REGION Network 2: ADDRESS 2
   RUNG wire#powerrail
      { S7_Templates := "SrcType := Real"; S7_GenerateENO := "TRUE" } Div(in1 := "DB6_MAV2_DBD".ADDRES_2, in2 := 32.768, out => "DB6_MAV2_DBD".SCALLING_2)
      { S7_Templates := "[SrcType := Real, DestType := DInt]"; S7_GenerateENO := "TRUE" } Round(in := "DB6_MAV2_DBD".SCALLING_2, out => "DB6_MAV2_DBD".STAT58)
      { S7_GenerateENO := "TRUE" } Move(in := "DB6_MAV2_DBD".STAT58, out1 => "DB7".STAT0)
   END_RUNG
   // the same network as SCL:
   // ENO of a box is taken as its EN; it also drops when the box reports an error
   "DB6_MAV2_DBD".SCALLING_2 := "DB6_MAV2_DBD".ADDRES_2 / 32.768;
   "DB6_MAV2_DBD".STAT58 := ROUND("DB6_MAV2_DBD".SCALLING_2);
   "DB7".STAT0 := "DB6_MAV2_DBD".STAT58;
END_REGION

REGION Network 3: ADDRESS 3
   RUNG wire#powerrail
      { S7_Templates := "[SrcType := Int, DestType := DInt]"; S7_GenerateENO := "TRUE" } Convert(in := "DB5_MAV".ADDRES_3, out => "DB8_SCALLING_MAV".ADDRESS_3)
      { S7_Templates := "[SrcType := DInt, DestType := Real]"; S7_GenerateENO := "TRUE" } Convert(in := "DB8_SCALLING_MAV".ADDRESS_3, out => "DB6_MAV2_DBD".ADDRES_3)
   END_RUNG
   // the same network as SCL:
   // ENO of a box is taken as its EN; it also drops when the box reports an error
   "DB8_SCALLING_MAV".ADDRESS_3 := INT_TO_DINT("DB5_MAV".ADDRES_3);
   "DB6_MAV2_DBD".ADDRES_3 := DINT_TO_REAL("DB8_SCALLING_MAV".ADDRESS_3);
END_REGION

REGION Network 4: ADDRESS 3
   RUNG wire#powerrail
      { S7_Templates := "SrcType := Real"; S7_GenerateENO := "TRUE" } Div(in1 := "DB6_MAV2_DBD".ADDRES_3, in2 := 32.768, out => "DB6_MAV2_DBD".SCALLING_3)
      { S7_Templates := "[SrcType := Real, DestType := DInt]"; S7_GenerateENO := "TRUE" } Round(in := "DB6_MAV2_DBD".SCALLING_3, out => "DB6_MAV2_DBD".STAT59)
      { S7_GenerateENO := "TRUE" } Move(in := "DB6_MAV2_DBD".STAT59, out1 => "DB7".STAT1)
   END_RUNG
   // the same network as SCL:
   // ENO of a box is taken as its EN; it also drops when the box reports an error
   "DB6_MAV2_DBD".SCALLING_3 := "DB6_MAV2_DBD".ADDRES_3 / 32.768;
   "DB6_MAV2_DBD".STAT59 := ROUND("DB6_MAV2_DBD".SCALLING_3);
   "DB7".STAT1 := "DB6_MAV2_DBD".STAT59;
END_REGION

REGION Network 5: ADDRESS 4
   RUNG wire#powerrail
      { S7_Templates := "[SrcType := Int, DestType := DInt]"; S7_GenerateENO := "TRUE" } Convert(in := "DB5_MAV".ADDRES_4, out => "DB8_SCALLING_MAV".ADDRESS_4)
      { S7_Templates := "[SrcType := DInt, DestType := Real]"; S7_GenerateENO := "TRUE" } Convert(in := "DB8_SCALLING_MAV".ADDRESS_4, out => "DB6_MAV2_DBD".ADDRES_4)
   END_RUNG
   // the same network as SCL:
   // ENO of a box is taken as its EN; it also drops when the box reports an error
   "DB8_SCALLING_MAV".ADDRESS_4 := INT_TO_DINT("DB5_MAV".ADDRES_4);
   "DB6_MAV2_DBD".ADDRES_4 := DINT_TO_REAL("DB8_SCALLING_MAV".ADDRESS_4);
END_REGION

REGION Network 6: ADDRESS 4
   RUNG wire#powerrail
      { S7_Templates := "SrcType := Real"; S7_GenerateENO := "TRUE" } Div(in1 := "DB6_MAV2_DBD".ADDRES_4, in2 := 32.768, out => "DB6_MAV2_DBD".SCALLING_4)
      { S7_Templates := "[SrcType := Real, DestType := DInt]"; S7_GenerateENO := "TRUE" } Round(in := "DB6_MAV2_DBD".SCALLING_4, out => "DB6_MAV2_DBD".STAT60)
      { S7_GenerateENO := "TRUE" } Move(in := "DB6_MAV2_DBD".STAT60, out1 => "DB7".STAT2)
   END_RUNG
   // the same network as SCL:
   // ENO of a box is taken as its EN; it also drops when the box reports an error
   "DB6_MAV2_DBD".SCALLING_4 := "DB6_MAV2_DBD".ADDRES_4 / 32.768;
   "DB6_MAV2_DBD".STAT60 := ROUND("DB6_MAV2_DBD".SCALLING_4);
   "DB7".STAT2 := "DB6_MAV2_DBD".STAT60;
END_REGION

REGION Network 7: ADDRESS 5
   RUNG wire#powerrail
      { S7_Templates := "[SrcType := Int, DestType := DInt]"; S7_GenerateENO := "TRUE" } Convert(in := "DB5_MAV".ADDRES_5, out => "DB8_SCALLING_MAV".ADDRESS_5)
      { S7_Templates := "[SrcType := DInt, DestType := Real]"; S7_GenerateENO := "TRUE" } Convert(in := "DB8_SCALLING_MAV".ADDRESS_5, out => "DB6_MAV2_DBD".ADDRES_5)
   END_RUNG
   // the same network as SCL:
   // ENO of a box is taken as its EN; it also drops when the box reports an error
   "DB8_SCALLING_MAV".ADDRESS_5 := INT_TO_DINT("DB5_MAV".ADDRES_5);
   "DB6_MAV2_DBD".ADDRES_5 := DINT_TO_REAL("DB8_SCALLING_MAV".ADDRESS_5);
END_REGION

REGION Network 8: ADDRESS 5
   RUNG wire#powerrail
      { S7_Templates := "SrcType := Real"; S7_GenerateENO := "TRUE" } Div(in1 := "DB6_MAV2_DBD".ADDRES_5, in2 := 32.768, out => "DB6_MAV2_DBD".SCALLING_5)
      { S7_Templates := "[SrcType := Real, DestType := DInt]"; S7_GenerateENO := "TRUE" } Round(in := "DB6_MAV2_DBD".SCALLING_5, out => "DB6_MAV2_DBD".STAT61)
      { S7_GenerateENO := "TRUE" } Move(in := "DB6_MAV2_DBD".STAT61, out1 => "DB7".STAT3)
   END_RUNG
   // the same network as SCL:
   // ENO of a box is taken as its EN; it also drops when the box reports an error
   "DB6_MAV2_DBD".SCALLING_5 := "DB6_MAV2_DBD".ADDRES_5 / 32.768;
   "DB6_MAV2_DBD".STAT61 := ROUND("DB6_MAV2_DBD".SCALLING_5);
   "DB7".STAT3 := "DB6_MAV2_DBD".STAT61;
END_REGION

REGION Network 9: ADDRESS 6
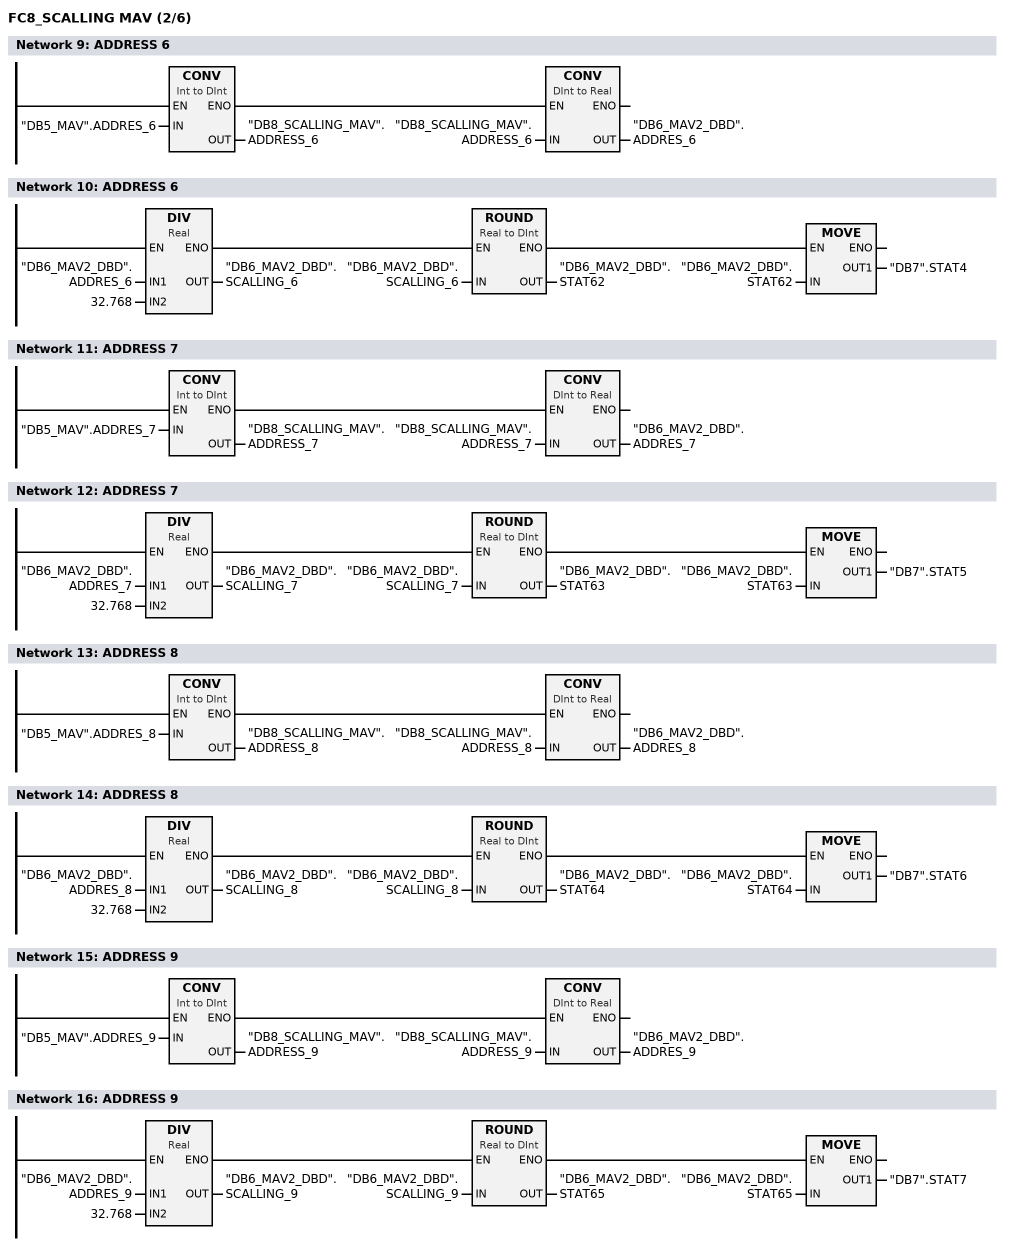
   RUNG wire#powerrail
      { S7_Templates := "[SrcType := Int, DestType := DInt]"; S7_GenerateENO := "TRUE" } Convert(in := "DB5_MAV".ADDRES_6, out => "DB8_SCALLING_MAV".ADDRESS_6)
      { S7_Templates := "[SrcType := DInt, DestType := Real]"; S7_GenerateENO := "TRUE" } Convert(in := "DB8_SCALLING_MAV".ADDRESS_6, out => "DB6_MAV2_DBD".ADDRES_6)
   END_RUNG
   // the same network as SCL:
   // ENO of a box is taken as its EN; it also drops when the box reports an error
   "DB8_SCALLING_MAV".ADDRESS_6 := INT_TO_DINT("DB5_MAV".ADDRES_6);
   "DB6_MAV2_DBD".ADDRES_6 := DINT_TO_REAL("DB8_SCALLING_MAV".ADDRESS_6);
END_REGION

REGION Network 10: ADDRESS 6
   RUNG wire#powerrail
      { S7_Templates := "SrcType := Real"; S7_GenerateENO := "TRUE" } Div(in1 := "DB6_MAV2_DBD".ADDRES_6, in2 := 32.768, out => "DB6_MAV2_DBD".SCALLING_6)
      { S7_Templates := "[SrcType := Real, DestType := DInt]"; S7_GenerateENO := "TRUE" } Round(in := "DB6_MAV2_DBD".SCALLING_6, out => "DB6_MAV2_DBD".STAT62)
      { S7_GenerateENO := "TRUE" } Move(in := "DB6_MAV2_DBD".STAT62, out1 => "DB7".STAT4)
   END_RUNG
   // the same network as SCL:
   // ENO of a box is taken as its EN; it also drops when the box reports an error
   "DB6_MAV2_DBD".SCALLING_6 := "DB6_MAV2_DBD".ADDRES_6 / 32.768;
   "DB6_MAV2_DBD".STAT62 := ROUND("DB6_MAV2_DBD".SCALLING_6);
   "DB7".STAT4 := "DB6_MAV2_DBD".STAT62;
END_REGION

REGION Network 11: ADDRESS 7
   RUNG wire#powerrail
      { S7_Templates := "[SrcType := Int, DestType := DInt]"; S7_GenerateENO := "TRUE" } Convert(in := "DB5_MAV".ADDRES_7, out => "DB8_SCALLING_MAV".ADDRESS_7)
      { S7_Templates := "[SrcType := DInt, DestType := Real]"; S7_GenerateENO := "TRUE" } Convert(in := "DB8_SCALLING_MAV".ADDRESS_7, out => "DB6_MAV2_DBD".ADDRES_7)
   END_RUNG
   // the same network as SCL:
   // ENO of a box is taken as its EN; it also drops when the box reports an error
   "DB8_SCALLING_MAV".ADDRESS_7 := INT_TO_DINT("DB5_MAV".ADDRES_7);
   "DB6_MAV2_DBD".ADDRES_7 := DINT_TO_REAL("DB8_SCALLING_MAV".ADDRESS_7);
END_REGION

REGION Network 12: ADDRESS 7
   RUNG wire#powerrail
      { S7_Templates := "SrcType := Real"; S7_GenerateENO := "TRUE" } Div(in1 := "DB6_MAV2_DBD".ADDRES_7, in2 := 32.768, out => "DB6_MAV2_DBD".SCALLING_7)
      { S7_Templates := "[SrcType := Real, DestType := DInt]"; S7_GenerateENO := "TRUE" } Round(in := "DB6_MAV2_DBD".SCALLING_7, out => "DB6_MAV2_DBD".STAT63)
      { S7_GenerateENO := "TRUE" } Move(in := "DB6_MAV2_DBD".STAT63, out1 => "DB7".STAT5)
   END_RUNG
   // the same network as SCL:
   // ENO of a box is taken as its EN; it also drops when the box reports an error
   "DB6_MAV2_DBD".SCALLING_7 := "DB6_MAV2_DBD".ADDRES_7 / 32.768;
   "DB6_MAV2_DBD".STAT63 := ROUND("DB6_MAV2_DBD".SCALLING_7);
   "DB7".STAT5 := "DB6_MAV2_DBD".STAT63;
END_REGION

REGION Network 13: ADDRESS 8
   RUNG wire#powerrail
      { S7_Templates := "[SrcType := Int, DestType := DInt]"; S7_GenerateENO := "TRUE" } Convert(in := "DB5_MAV".ADDRES_8, out => "DB8_SCALLING_MAV".ADDRESS_8)
      { S7_Templates := "[SrcType := DInt, DestType := Real]"; S7_GenerateENO := "TRUE" } Convert(in := "DB8_SCALLING_MAV".ADDRESS_8, out => "DB6_MAV2_DBD".ADDRES_8)
   END_RUNG
   // the same network as SCL:
   // ENO of a box is taken as its EN; it also drops when the box reports an error
   "DB8_SCALLING_MAV".ADDRESS_8 := INT_TO_DINT("DB5_MAV".ADDRES_8);
   "DB6_MAV2_DBD".ADDRES_8 := DINT_TO_REAL("DB8_SCALLING_MAV".ADDRESS_8);
END_REGION

REGION Network 14: ADDRESS 8
   RUNG wire#powerrail
      { S7_Templates := "SrcType := Real"; S7_GenerateENO := "TRUE" } Div(in1 := "DB6_MAV2_DBD".ADDRES_8, in2 := 32.768, out => "DB6_MAV2_DBD".SCALLING_8)
      { S7_Templates := "[SrcType := Real, DestType := DInt]"; S7_GenerateENO := "TRUE" } Round(in := "DB6_MAV2_DBD".SCALLING_8, out => "DB6_MAV2_DBD".STAT64)
      { S7_GenerateENO := "TRUE" } Move(in := "DB6_MAV2_DBD".STAT64, out1 => "DB7".STAT6)
   END_RUNG
   // the same network as SCL:
   // ENO of a box is taken as its EN; it also drops when the box reports an error
   "DB6_MAV2_DBD".SCALLING_8 := "DB6_MAV2_DBD".ADDRES_8 / 32.768;
   "DB6_MAV2_DBD".STAT64 := ROUND("DB6_MAV2_DBD".SCALLING_8);
   "DB7".STAT6 := "DB6_MAV2_DBD".STAT64;
END_REGION

REGION Network 15: ADDRESS 9
   RUNG wire#powerrail
      { S7_Templates := "[SrcType := Int, DestType := DInt]"; S7_GenerateENO := "TRUE" } Convert(in := "DB5_MAV".ADDRES_9, out => "DB8_SCALLING_MAV".ADDRESS_9)
      { S7_Templates := "[SrcType := DInt, DestType := Real]"; S7_GenerateENO := "TRUE" } Convert(in := "DB8_SCALLING_MAV".ADDRESS_9, out => "DB6_MAV2_DBD".ADDRES_9)
   END_RUNG
   // the same network as SCL:
   // ENO of a box is taken as its EN; it also drops when the box reports an error
   "DB8_SCALLING_MAV".ADDRESS_9 := INT_TO_DINT("DB5_MAV".ADDRES_9);
   "DB6_MAV2_DBD".ADDRES_9 := DINT_TO_REAL("DB8_SCALLING_MAV".ADDRESS_9);
END_REGION

REGION Network 16: ADDRESS 9
   RUNG wire#powerrail
      { S7_Templates := "SrcType := Real"; S7_GenerateENO := "TRUE" } Div(in1 := "DB6_MAV2_DBD".ADDRES_9, in2 := 32.768, out => "DB6_MAV2_DBD".SCALLING_9)
      { S7_Templates := "[SrcType := Real, DestType := DInt]"; S7_GenerateENO := "TRUE" } Round(in := "DB6_MAV2_DBD".SCALLING_9, out => "DB6_MAV2_DBD".STAT65)
      { S7_GenerateENO := "TRUE" } Move(in := "DB6_MAV2_DBD".STAT65, out1 => "DB7".STAT7)
   END_RUNG
   // the same network as SCL:
   // ENO of a box is taken as its EN; it also drops when the box reports an error
   "DB6_MAV2_DBD".SCALLING_9 := "DB6_MAV2_DBD".ADDRES_9 / 32.768;
   "DB6_MAV2_DBD".STAT65 := ROUND("DB6_MAV2_DBD".SCALLING_9);
   "DB7".STAT7 := "DB6_MAV2_DBD".STAT65;
END_REGION

REGION Network 17: ADDRESS 10
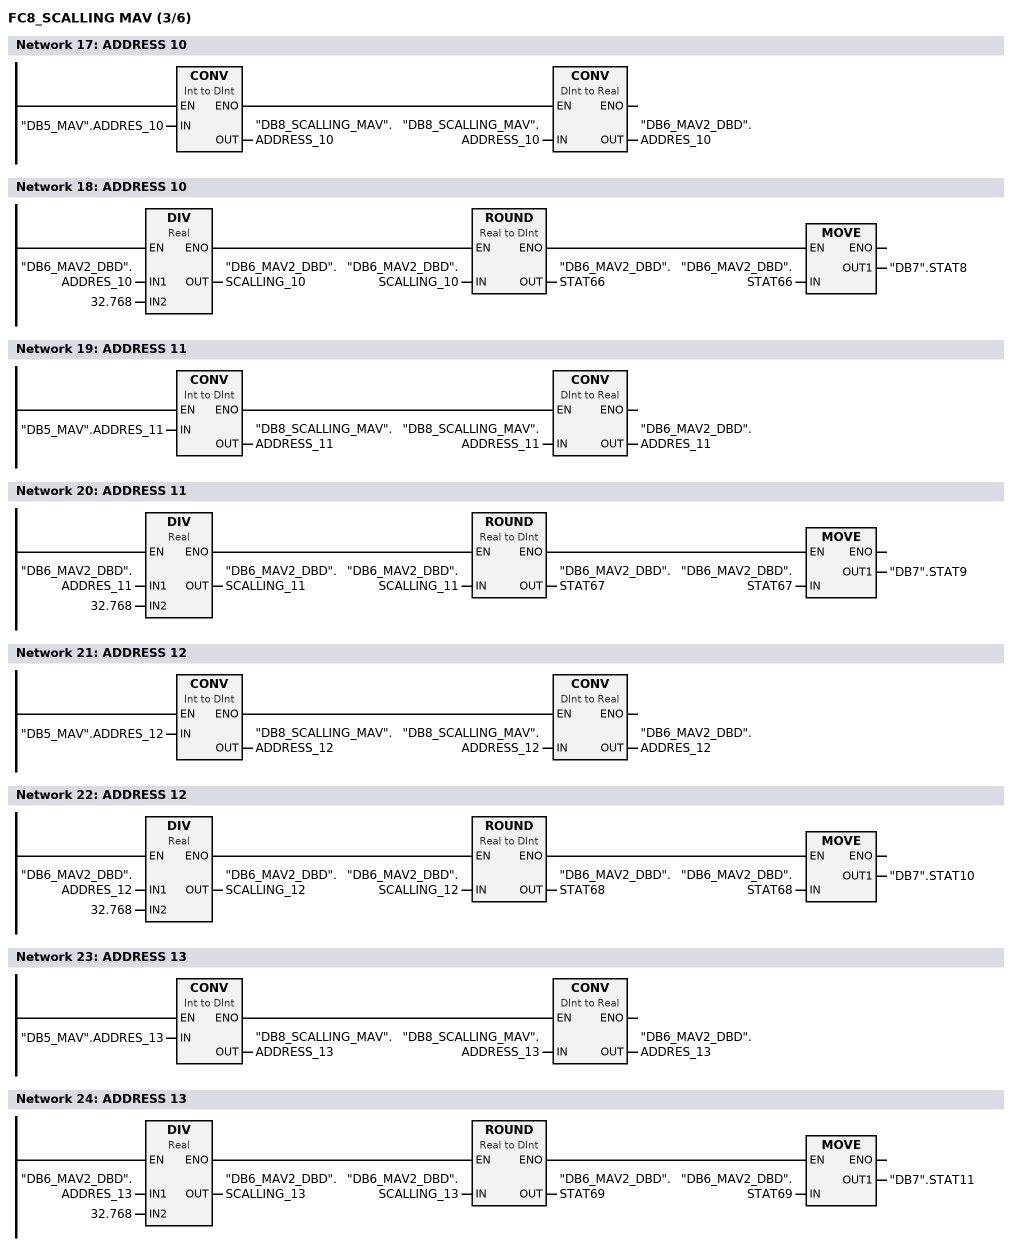
   RUNG wire#powerrail
      { S7_Templates := "[SrcType := Int, DestType := DInt]"; S7_GenerateENO := "TRUE" } Convert(in := "DB5_MAV".ADDRES_10, out => "DB8_SCALLING_MAV".ADDRESS_10)
      { S7_Templates := "[SrcType := DInt, DestType := Real]"; S7_GenerateENO := "TRUE" } Convert(in := "DB8_SCALLING_MAV".ADDRESS_10, out => "DB6_MAV2_DBD".ADDRES_10)
   END_RUNG
   // the same network as SCL:
   // ENO of a box is taken as its EN; it also drops when the box reports an error
   "DB8_SCALLING_MAV".ADDRESS_10 := INT_TO_DINT("DB5_MAV".ADDRES_10);
   "DB6_MAV2_DBD".ADDRES_10 := DINT_TO_REAL("DB8_SCALLING_MAV".ADDRESS_10);
END_REGION

REGION Network 18: ADDRESS 10
   RUNG wire#powerrail
      { S7_Templates := "SrcType := Real"; S7_GenerateENO := "TRUE" } Div(in1 := "DB6_MAV2_DBD".ADDRES_10, in2 := 32.768, out => "DB6_MAV2_DBD".SCALLING_10)
      { S7_Templates := "[SrcType := Real, DestType := DInt]"; S7_GenerateENO := "TRUE" } Round(in := "DB6_MAV2_DBD".SCALLING_10, out => "DB6_MAV2_DBD".STAT66)
      { S7_GenerateENO := "TRUE" } Move(in := "DB6_MAV2_DBD".STAT66, out1 => "DB7".STAT8)
   END_RUNG
   // the same network as SCL:
   // ENO of a box is taken as its EN; it also drops when the box reports an error
   "DB6_MAV2_DBD".SCALLING_10 := "DB6_MAV2_DBD".ADDRES_10 / 32.768;
   "DB6_MAV2_DBD".STAT66 := ROUND("DB6_MAV2_DBD".SCALLING_10);
   "DB7".STAT8 := "DB6_MAV2_DBD".STAT66;
END_REGION

REGION Network 19: ADDRESS 11
   RUNG wire#powerrail
      { S7_Templates := "[SrcType := Int, DestType := DInt]"; S7_GenerateENO := "TRUE" } Convert(in := "DB5_MAV".ADDRES_11, out => "DB8_SCALLING_MAV".ADDRESS_11)
      { S7_Templates := "[SrcType := DInt, DestType := Real]"; S7_GenerateENO := "TRUE" } Convert(in := "DB8_SCALLING_MAV".ADDRESS_11, out => "DB6_MAV2_DBD".ADDRES_11)
   END_RUNG
   // the same network as SCL:
   // ENO of a box is taken as its EN; it also drops when the box reports an error
   "DB8_SCALLING_MAV".ADDRESS_11 := INT_TO_DINT("DB5_MAV".ADDRES_11);
   "DB6_MAV2_DBD".ADDRES_11 := DINT_TO_REAL("DB8_SCALLING_MAV".ADDRESS_11);
END_REGION

REGION Network 20: ADDRESS 11
   RUNG wire#powerrail
      { S7_Templates := "SrcType := Real"; S7_GenerateENO := "TRUE" } Div(in1 := "DB6_MAV2_DBD".ADDRES_11, in2 := 32.768, out => "DB6_MAV2_DBD".SCALLING_11)
      { S7_Templates := "[SrcType := Real, DestType := DInt]"; S7_GenerateENO := "TRUE" } Round(in := "DB6_MAV2_DBD".SCALLING_11, out => "DB6_MAV2_DBD".STAT67)
      { S7_GenerateENO := "TRUE" } Move(in := "DB6_MAV2_DBD".STAT67, out1 => "DB7".STAT9)
   END_RUNG
   // the same network as SCL:
   // ENO of a box is taken as its EN; it also drops when the box reports an error
   "DB6_MAV2_DBD".SCALLING_11 := "DB6_MAV2_DBD".ADDRES_11 / 32.768;
   "DB6_MAV2_DBD".STAT67 := ROUND("DB6_MAV2_DBD".SCALLING_11);
   "DB7".STAT9 := "DB6_MAV2_DBD".STAT67;
END_REGION

REGION Network 21: ADDRESS 12
   RUNG wire#powerrail
      { S7_Templates := "[SrcType := Int, DestType := DInt]"; S7_GenerateENO := "TRUE" } Convert(in := "DB5_MAV".ADDRES_12, out => "DB8_SCALLING_MAV".ADDRESS_12)
      { S7_Templates := "[SrcType := DInt, DestType := Real]"; S7_GenerateENO := "TRUE" } Convert(in := "DB8_SCALLING_MAV".ADDRESS_12, out => "DB6_MAV2_DBD".ADDRES_12)
   END_RUNG
   // the same network as SCL:
   // ENO of a box is taken as its EN; it also drops when the box reports an error
   "DB8_SCALLING_MAV".ADDRESS_12 := INT_TO_DINT("DB5_MAV".ADDRES_12);
   "DB6_MAV2_DBD".ADDRES_12 := DINT_TO_REAL("DB8_SCALLING_MAV".ADDRESS_12);
END_REGION

REGION Network 22: ADDRESS 12
   RUNG wire#powerrail
      { S7_Templates := "SrcType := Real"; S7_GenerateENO := "TRUE" } Div(in1 := "DB6_MAV2_DBD".ADDRES_12, in2 := 32.768, out => "DB6_MAV2_DBD".SCALLING_12)
      { S7_Templates := "[SrcType := Real, DestType := DInt]"; S7_GenerateENO := "TRUE" } Round(in := "DB6_MAV2_DBD".SCALLING_12, out => "DB6_MAV2_DBD".STAT68)
      { S7_GenerateENO := "TRUE" } Move(in := "DB6_MAV2_DBD".STAT68, out1 => "DB7".STAT10)
   END_RUNG
   // the same network as SCL:
   // ENO of a box is taken as its EN; it also drops when the box reports an error
   "DB6_MAV2_DBD".SCALLING_12 := "DB6_MAV2_DBD".ADDRES_12 / 32.768;
   "DB6_MAV2_DBD".STAT68 := ROUND("DB6_MAV2_DBD".SCALLING_12);
   "DB7".STAT10 := "DB6_MAV2_DBD".STAT68;
END_REGION

REGION Network 23: ADDRESS 13
   RUNG wire#powerrail
      { S7_Templates := "[SrcType := Int, DestType := DInt]"; S7_GenerateENO := "TRUE" } Convert(in := "DB5_MAV".ADDRES_13, out => "DB8_SCALLING_MAV".ADDRESS_13)
      { S7_Templates := "[SrcType := DInt, DestType := Real]"; S7_GenerateENO := "TRUE" } Convert(in := "DB8_SCALLING_MAV".ADDRESS_13, out => "DB6_MAV2_DBD".ADDRES_13)
   END_RUNG
   // the same network as SCL:
   // ENO of a box is taken as its EN; it also drops when the box reports an error
   "DB8_SCALLING_MAV".ADDRESS_13 := INT_TO_DINT("DB5_MAV".ADDRES_13);
   "DB6_MAV2_DBD".ADDRES_13 := DINT_TO_REAL("DB8_SCALLING_MAV".ADDRESS_13);
END_REGION

REGION Network 24: ADDRESS 13
   RUNG wire#powerrail
      { S7_Templates := "SrcType := Real"; S7_GenerateENO := "TRUE" } Div(in1 := "DB6_MAV2_DBD".ADDRES_13, in2 := 32.768, out => "DB6_MAV2_DBD".SCALLING_13)
      { S7_Templates := "[SrcType := Real, DestType := DInt]"; S7_GenerateENO := "TRUE" } Round(in := "DB6_MAV2_DBD".SCALLING_13, out => "DB6_MAV2_DBD".STAT69)
      { S7_GenerateENO := "TRUE" } Move(in := "DB6_MAV2_DBD".STAT69, out1 => "DB7".STAT11)
   END_RUNG
   // the same network as SCL:
   // ENO of a box is taken as its EN; it also drops when the box reports an error
   "DB6_MAV2_DBD".SCALLING_13 := "DB6_MAV2_DBD".ADDRES_13 / 32.768;
   "DB6_MAV2_DBD".STAT69 := ROUND("DB6_MAV2_DBD".SCALLING_13);
   "DB7".STAT11 := "DB6_MAV2_DBD".STAT69;
END_REGION

REGION Network 25: ADDRESS 14
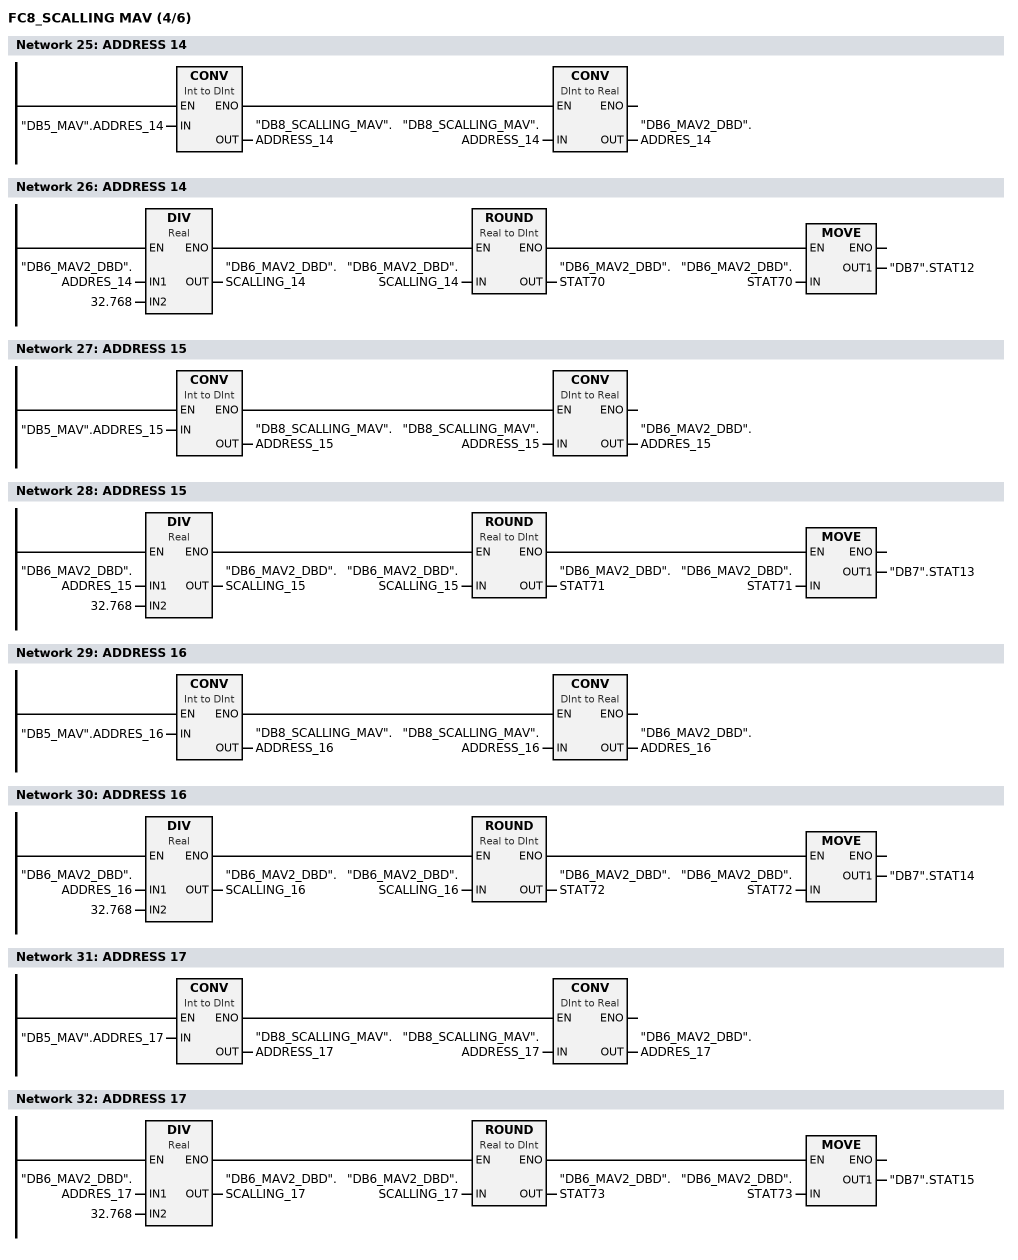
   RUNG wire#powerrail
      { S7_Templates := "[SrcType := Int, DestType := DInt]"; S7_GenerateENO := "TRUE" } Convert(in := "DB5_MAV".ADDRES_14, out => "DB8_SCALLING_MAV".ADDRESS_14)
      { S7_Templates := "[SrcType := DInt, DestType := Real]"; S7_GenerateENO := "TRUE" } Convert(in := "DB8_SCALLING_MAV".ADDRESS_14, out => "DB6_MAV2_DBD".ADDRES_14)
   END_RUNG
   // the same network as SCL:
   // ENO of a box is taken as its EN; it also drops when the box reports an error
   "DB8_SCALLING_MAV".ADDRESS_14 := INT_TO_DINT("DB5_MAV".ADDRES_14);
   "DB6_MAV2_DBD".ADDRES_14 := DINT_TO_REAL("DB8_SCALLING_MAV".ADDRESS_14);
END_REGION

REGION Network 26: ADDRESS 14
   RUNG wire#powerrail
      { S7_Templates := "SrcType := Real"; S7_GenerateENO := "TRUE" } Div(in1 := "DB6_MAV2_DBD".ADDRES_14, in2 := 32.768, out => "DB6_MAV2_DBD".SCALLING_14)
      { S7_Templates := "[SrcType := Real, DestType := DInt]"; S7_GenerateENO := "TRUE" } Round(in := "DB6_MAV2_DBD".SCALLING_14, out => "DB6_MAV2_DBD".STAT70)
      { S7_GenerateENO := "TRUE" } Move(in := "DB6_MAV2_DBD".STAT70, out1 => "DB7".STAT12)
   END_RUNG
   // the same network as SCL:
   // ENO of a box is taken as its EN; it also drops when the box reports an error
   "DB6_MAV2_DBD".SCALLING_14 := "DB6_MAV2_DBD".ADDRES_14 / 32.768;
   "DB6_MAV2_DBD".STAT70 := ROUND("DB6_MAV2_DBD".SCALLING_14);
   "DB7".STAT12 := "DB6_MAV2_DBD".STAT70;
END_REGION

REGION Network 27: ADDRESS 15
   RUNG wire#powerrail
      { S7_Templates := "[SrcType := Int, DestType := DInt]"; S7_GenerateENO := "TRUE" } Convert(in := "DB5_MAV".ADDRES_15, out => "DB8_SCALLING_MAV".ADDRESS_15)
      { S7_Templates := "[SrcType := DInt, DestType := Real]"; S7_GenerateENO := "TRUE" } Convert(in := "DB8_SCALLING_MAV".ADDRESS_15, out => "DB6_MAV2_DBD".ADDRES_15)
   END_RUNG
   // the same network as SCL:
   // ENO of a box is taken as its EN; it also drops when the box reports an error
   "DB8_SCALLING_MAV".ADDRESS_15 := INT_TO_DINT("DB5_MAV".ADDRES_15);
   "DB6_MAV2_DBD".ADDRES_15 := DINT_TO_REAL("DB8_SCALLING_MAV".ADDRESS_15);
END_REGION

REGION Network 28: ADDRESS 15
   RUNG wire#powerrail
      { S7_Templates := "SrcType := Real"; S7_GenerateENO := "TRUE" } Div(in1 := "DB6_MAV2_DBD".ADDRES_15, in2 := 32.768, out => "DB6_MAV2_DBD".SCALLING_15)
      { S7_Templates := "[SrcType := Real, DestType := DInt]"; S7_GenerateENO := "TRUE" } Round(in := "DB6_MAV2_DBD".SCALLING_15, out => "DB6_MAV2_DBD".STAT71)
      { S7_GenerateENO := "TRUE" } Move(in := "DB6_MAV2_DBD".STAT71, out1 => "DB7".STAT13)
   END_RUNG
   // the same network as SCL:
   // ENO of a box is taken as its EN; it also drops when the box reports an error
   "DB6_MAV2_DBD".SCALLING_15 := "DB6_MAV2_DBD".ADDRES_15 / 32.768;
   "DB6_MAV2_DBD".STAT71 := ROUND("DB6_MAV2_DBD".SCALLING_15);
   "DB7".STAT13 := "DB6_MAV2_DBD".STAT71;
END_REGION

REGION Network 29: ADDRESS 16
   RUNG wire#powerrail
      { S7_Templates := "[SrcType := Int, DestType := DInt]"; S7_GenerateENO := "TRUE" } Convert(in := "DB5_MAV".ADDRES_16, out => "DB8_SCALLING_MAV".ADDRESS_16)
      { S7_Templates := "[SrcType := DInt, DestType := Real]"; S7_GenerateENO := "TRUE" } Convert(in := "DB8_SCALLING_MAV".ADDRESS_16, out => "DB6_MAV2_DBD".ADDRES_16)
   END_RUNG
   // the same network as SCL:
   // ENO of a box is taken as its EN; it also drops when the box reports an error
   "DB8_SCALLING_MAV".ADDRESS_16 := INT_TO_DINT("DB5_MAV".ADDRES_16);
   "DB6_MAV2_DBD".ADDRES_16 := DINT_TO_REAL("DB8_SCALLING_MAV".ADDRESS_16);
END_REGION

REGION Network 30: ADDRESS 16
   RUNG wire#powerrail
      { S7_Templates := "SrcType := Real"; S7_GenerateENO := "TRUE" } Div(in1 := "DB6_MAV2_DBD".ADDRES_16, in2 := 32.768, out => "DB6_MAV2_DBD".SCALLING_16)
      { S7_Templates := "[SrcType := Real, DestType := DInt]"; S7_GenerateENO := "TRUE" } Round(in := "DB6_MAV2_DBD".SCALLING_16, out => "DB6_MAV2_DBD".STAT72)
      { S7_GenerateENO := "TRUE" } Move(in := "DB6_MAV2_DBD".STAT72, out1 => "DB7".STAT14)
   END_RUNG
   // the same network as SCL:
   // ENO of a box is taken as its EN; it also drops when the box reports an error
   "DB6_MAV2_DBD".SCALLING_16 := "DB6_MAV2_DBD".ADDRES_16 / 32.768;
   "DB6_MAV2_DBD".STAT72 := ROUND("DB6_MAV2_DBD".SCALLING_16);
   "DB7".STAT14 := "DB6_MAV2_DBD".STAT72;
END_REGION

REGION Network 31: ADDRESS 17
   RUNG wire#powerrail
      { S7_Templates := "[SrcType := Int, DestType := DInt]"; S7_GenerateENO := "TRUE" } Convert(in := "DB5_MAV".ADDRES_17, out => "DB8_SCALLING_MAV".ADDRESS_17)
      { S7_Templates := "[SrcType := DInt, DestType := Real]"; S7_GenerateENO := "TRUE" } Convert(in := "DB8_SCALLING_MAV".ADDRESS_17, out => "DB6_MAV2_DBD".ADDRES_17)
   END_RUNG
   // the same network as SCL:
   // ENO of a box is taken as its EN; it also drops when the box reports an error
   "DB8_SCALLING_MAV".ADDRESS_17 := INT_TO_DINT("DB5_MAV".ADDRES_17);
   "DB6_MAV2_DBD".ADDRES_17 := DINT_TO_REAL("DB8_SCALLING_MAV".ADDRESS_17);
END_REGION

REGION Network 32: ADDRESS 17
   RUNG wire#powerrail
      { S7_Templates := "SrcType := Real"; S7_GenerateENO := "TRUE" } Div(in1 := "DB6_MAV2_DBD".ADDRES_17, in2 := 32.768, out => "DB6_MAV2_DBD".SCALLING_17)
      { S7_Templates := "[SrcType := Real, DestType := DInt]"; S7_GenerateENO := "TRUE" } Round(in := "DB6_MAV2_DBD".SCALLING_17, out => "DB6_MAV2_DBD".STAT73)
      { S7_GenerateENO := "TRUE" } Move(in := "DB6_MAV2_DBD".STAT73, out1 => "DB7".STAT15)
   END_RUNG
   // the same network as SCL:
   // ENO of a box is taken as its EN; it also drops when the box reports an error
   "DB6_MAV2_DBD".SCALLING_17 := "DB6_MAV2_DBD".ADDRES_17 / 32.768;
   "DB6_MAV2_DBD".STAT73 := ROUND("DB6_MAV2_DBD".SCALLING_17);
   "DB7".STAT15 := "DB6_MAV2_DBD".STAT73;
END_REGION

REGION Network 33: ADDRESS 18
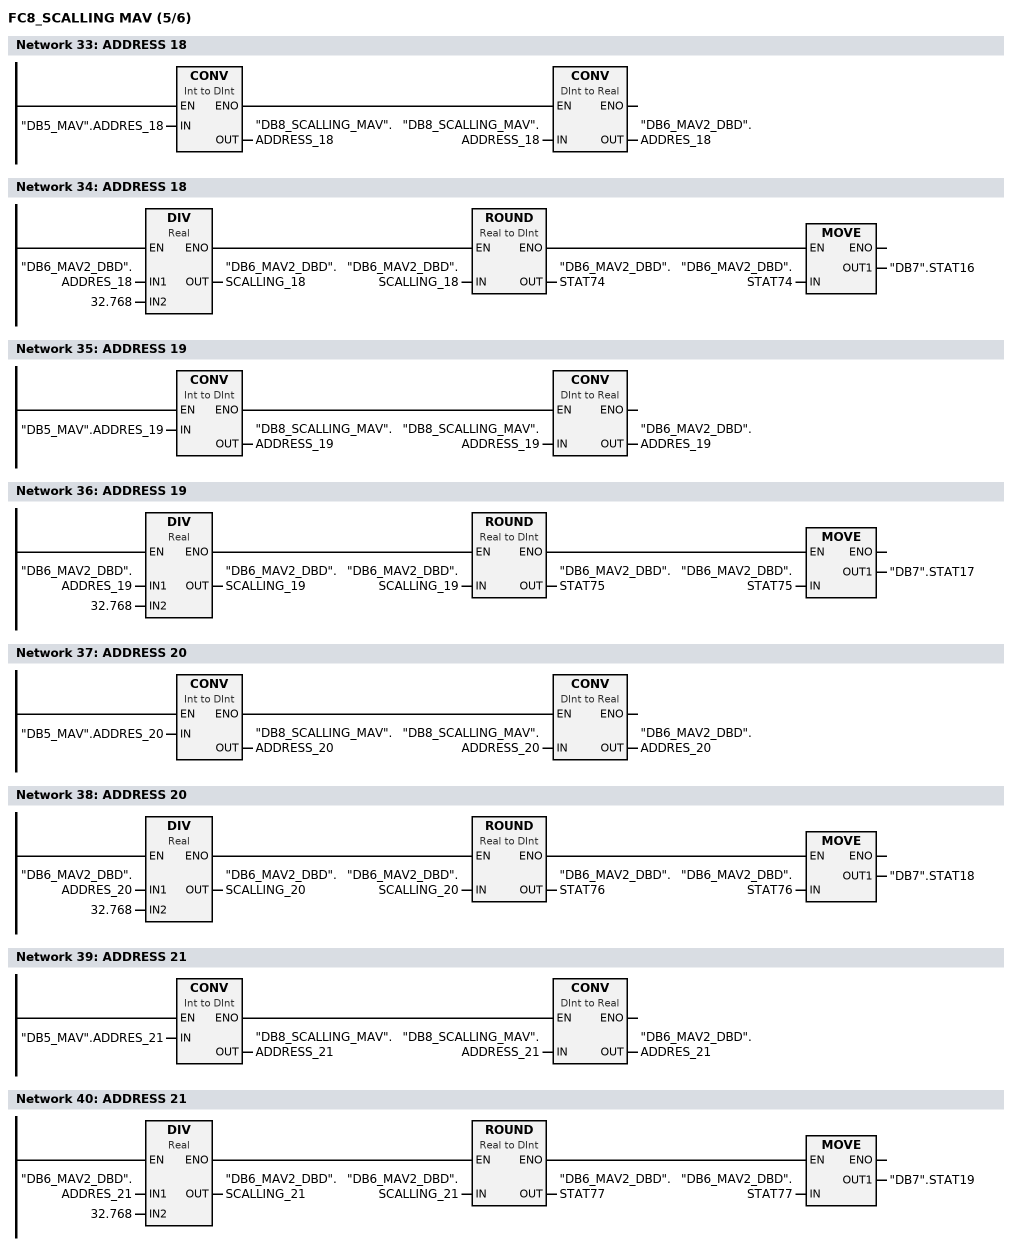
   RUNG wire#powerrail
      { S7_Templates := "[SrcType := Int, DestType := DInt]"; S7_GenerateENO := "TRUE" } Convert(in := "DB5_MAV".ADDRES_18, out => "DB8_SCALLING_MAV".ADDRESS_18)
      { S7_Templates := "[SrcType := DInt, DestType := Real]"; S7_GenerateENO := "TRUE" } Convert(in := "DB8_SCALLING_MAV".ADDRESS_18, out => "DB6_MAV2_DBD".ADDRES_18)
   END_RUNG
   // the same network as SCL:
   // ENO of a box is taken as its EN; it also drops when the box reports an error
   "DB8_SCALLING_MAV".ADDRESS_18 := INT_TO_DINT("DB5_MAV".ADDRES_18);
   "DB6_MAV2_DBD".ADDRES_18 := DINT_TO_REAL("DB8_SCALLING_MAV".ADDRESS_18);
END_REGION

REGION Network 34: ADDRESS 18
   RUNG wire#powerrail
      { S7_Templates := "SrcType := Real"; S7_GenerateENO := "TRUE" } Div(in1 := "DB6_MAV2_DBD".ADDRES_18, in2 := 32.768, out => "DB6_MAV2_DBD".SCALLING_18)
      { S7_Templates := "[SrcType := Real, DestType := DInt]"; S7_GenerateENO := "TRUE" } Round(in := "DB6_MAV2_DBD".SCALLING_18, out => "DB6_MAV2_DBD".STAT74)
      { S7_GenerateENO := "TRUE" } Move(in := "DB6_MAV2_DBD".STAT74, out1 => "DB7".STAT16)
   END_RUNG
   // the same network as SCL:
   // ENO of a box is taken as its EN; it also drops when the box reports an error
   "DB6_MAV2_DBD".SCALLING_18 := "DB6_MAV2_DBD".ADDRES_18 / 32.768;
   "DB6_MAV2_DBD".STAT74 := ROUND("DB6_MAV2_DBD".SCALLING_18);
   "DB7".STAT16 := "DB6_MAV2_DBD".STAT74;
END_REGION

REGION Network 35: ADDRESS 19
   RUNG wire#powerrail
      { S7_Templates := "[SrcType := Int, DestType := DInt]"; S7_GenerateENO := "TRUE" } Convert(in := "DB5_MAV".ADDRES_19, out => "DB8_SCALLING_MAV".ADDRESS_19)
      { S7_Templates := "[SrcType := DInt, DestType := Real]"; S7_GenerateENO := "TRUE" } Convert(in := "DB8_SCALLING_MAV".ADDRESS_19, out => "DB6_MAV2_DBD".ADDRES_19)
   END_RUNG
   // the same network as SCL:
   // ENO of a box is taken as its EN; it also drops when the box reports an error
   "DB8_SCALLING_MAV".ADDRESS_19 := INT_TO_DINT("DB5_MAV".ADDRES_19);
   "DB6_MAV2_DBD".ADDRES_19 := DINT_TO_REAL("DB8_SCALLING_MAV".ADDRESS_19);
END_REGION

REGION Network 36: ADDRESS 19
   RUNG wire#powerrail
      { S7_Templates := "SrcType := Real"; S7_GenerateENO := "TRUE" } Div(in1 := "DB6_MAV2_DBD".ADDRES_19, in2 := 32.768, out => "DB6_MAV2_DBD".SCALLING_19)
      { S7_Templates := "[SrcType := Real, DestType := DInt]"; S7_GenerateENO := "TRUE" } Round(in := "DB6_MAV2_DBD".SCALLING_19, out => "DB6_MAV2_DBD".STAT75)
      { S7_GenerateENO := "TRUE" } Move(in := "DB6_MAV2_DBD".STAT75, out1 => "DB7".STAT17)
   END_RUNG
   // the same network as SCL:
   // ENO of a box is taken as its EN; it also drops when the box reports an error
   "DB6_MAV2_DBD".SCALLING_19 := "DB6_MAV2_DBD".ADDRES_19 / 32.768;
   "DB6_MAV2_DBD".STAT75 := ROUND("DB6_MAV2_DBD".SCALLING_19);
   "DB7".STAT17 := "DB6_MAV2_DBD".STAT75;
END_REGION

REGION Network 37: ADDRESS 20
   RUNG wire#powerrail
      { S7_Templates := "[SrcType := Int, DestType := DInt]"; S7_GenerateENO := "TRUE" } Convert(in := "DB5_MAV".ADDRES_20, out => "DB8_SCALLING_MAV".ADDRESS_20)
      { S7_Templates := "[SrcType := DInt, DestType := Real]"; S7_GenerateENO := "TRUE" } Convert(in := "DB8_SCALLING_MAV".ADDRESS_20, out => "DB6_MAV2_DBD".ADDRES_20)
   END_RUNG
   // the same network as SCL:
   // ENO of a box is taken as its EN; it also drops when the box reports an error
   "DB8_SCALLING_MAV".ADDRESS_20 := INT_TO_DINT("DB5_MAV".ADDRES_20);
   "DB6_MAV2_DBD".ADDRES_20 := DINT_TO_REAL("DB8_SCALLING_MAV".ADDRESS_20);
END_REGION

REGION Network 38: ADDRESS 20
   RUNG wire#powerrail
      { S7_Templates := "SrcType := Real"; S7_GenerateENO := "TRUE" } Div(in1 := "DB6_MAV2_DBD".ADDRES_20, in2 := 32.768, out => "DB6_MAV2_DBD".SCALLING_20)
      { S7_Templates := "[SrcType := Real, DestType := DInt]"; S7_GenerateENO := "TRUE" } Round(in := "DB6_MAV2_DBD".SCALLING_20, out => "DB6_MAV2_DBD".STAT76)
      { S7_GenerateENO := "TRUE" } Move(in := "DB6_MAV2_DBD".STAT76, out1 => "DB7".STAT18)
   END_RUNG
   // the same network as SCL:
   // ENO of a box is taken as its EN; it also drops when the box reports an error
   "DB6_MAV2_DBD".SCALLING_20 := "DB6_MAV2_DBD".ADDRES_20 / 32.768;
   "DB6_MAV2_DBD".STAT76 := ROUND("DB6_MAV2_DBD".SCALLING_20);
   "DB7".STAT18 := "DB6_MAV2_DBD".STAT76;
END_REGION

REGION Network 39: ADDRESS 21
   RUNG wire#powerrail
      { S7_Templates := "[SrcType := Int, DestType := DInt]"; S7_GenerateENO := "TRUE" } Convert(in := "DB5_MAV".ADDRES_21, out => "DB8_SCALLING_MAV".ADDRESS_21)
      { S7_Templates := "[SrcType := DInt, DestType := Real]"; S7_GenerateENO := "TRUE" } Convert(in := "DB8_SCALLING_MAV".ADDRESS_21, out => "DB6_MAV2_DBD".ADDRES_21)
   END_RUNG
   // the same network as SCL:
   // ENO of a box is taken as its EN; it also drops when the box reports an error
   "DB8_SCALLING_MAV".ADDRESS_21 := INT_TO_DINT("DB5_MAV".ADDRES_21);
   "DB6_MAV2_DBD".ADDRES_21 := DINT_TO_REAL("DB8_SCALLING_MAV".ADDRESS_21);
END_REGION

REGION Network 40: ADDRESS 21
   RUNG wire#powerrail
      { S7_Templates := "SrcType := Real"; S7_GenerateENO := "TRUE" } Div(in1 := "DB6_MAV2_DBD".ADDRES_21, in2 := 32.768, out => "DB6_MAV2_DBD".SCALLING_21)
      { S7_Templates := "[SrcType := Real, DestType := DInt]"; S7_GenerateENO := "TRUE" } Round(in := "DB6_MAV2_DBD".SCALLING_21, out => "DB6_MAV2_DBD".STAT77)
      { S7_GenerateENO := "TRUE" } Move(in := "DB6_MAV2_DBD".STAT77, out1 => "DB7".STAT19)
   END_RUNG
   // the same network as SCL:
   // ENO of a box is taken as its EN; it also drops when the box reports an error
   "DB6_MAV2_DBD".SCALLING_21 := "DB6_MAV2_DBD".ADDRES_21 / 32.768;
   "DB6_MAV2_DBD".STAT77 := ROUND("DB6_MAV2_DBD".SCALLING_21);
   "DB7".STAT19 := "DB6_MAV2_DBD".STAT77;
END_REGION

REGION Network 41: ADDRESS 22